               3:
                   IF (("req23" OR "reqdown3") AND "proximity23") THEN
                       #elevator2next := 3;
                   ELSIF ("req22" OR "reqdown2") THEN
                       #elevator2next := 2;
                       #elevator2heading := 1;
                   ELSIF ("req21" OR "reqdown1") THEN
                       #elevator2next := 1;
                       #elevator2heading := 1;
                   ELSIF ("req20") THEN
                       #elevator2next := 0;
                       #elevator2heading := 1;
                   ELSIF ("requpgnd") THEN
                       "requpgnd" := FALSE;
                       "req20" := TRUE;
                       #elevator2next := 0;
                       #elevator2heading := 1;
                   ELSIF ("requp1") THEN
                       "requp1" := FALSE;
                       "req21" := TRUE;
                       #elevator2next := 1;
                       #elevator2heading := 1;
                   ELSIF ("requp2") THEN
                       "requp2" := FALSE;
                       "req22" := TRUE;
                       #elevator2next := 2;
                       #elevator2heading := 1;
                   ELSE
                       #elevator2heading := 0;
                   END_IF;
               4:
                   IF (("req24" OR "reqdown4") AND "proximity24") THEN
                       #elevator2next := 4;
                   ELSIF ("req23" OR "reqdown3") THEN
                       #elevator2next := 3;
                       #elevator2heading := 1;
                   ELSIF ("req22" OR "reqdown2") THEN
                       #elevator2next := 2;
                       #elevator2heading := 1;
                   ELSIF ("req21" OR "reqdown1") THEN
                       #elevator2next := 1;
                       #elevator2heading := 1;
                   ELSIF ("req20") THEN
                       #elevator2next := 0;
                       #elevator2heading := 1;
                   ELSIF ("requpgnd") THEN
                       "requpgnd" := FALSE;
                       "req20" := TRUE;
                       #elevator2next := 0;
                       #elevator2heading := 1;
                   ELSIF ("requp1") THEN
                       "requp1" := FALSE;
                       "req21" := TRUE;
                       #elevator2next := 1;
                       #elevator2heading := 1;
                   ELSIF ("requp2") THEN
                       "requp2" := FALSE;
                       "req22" := TRUE;
                       #elevator2next := 2;
                       #elevator2heading := 1;
                   ELSIF ("requp3") THEN
                       "requp3" := FALSE;
                       "req23" := TRUE;
                       #elevator2next := 3;
                       #elevator2heading := 1;
                   ELSE
                       #elevator2heading := 0;
                   END_IF;

               5:
                   IF (("req25" OR "reqdown5") AND "proximity25") THEN
                       #elevator2next := 5;
                   ELSIF ("req24" OR "reqdown4") THEN
                       #elevator2next := 4;
                       #elevator2heading := 1;
                   ELSIF ("req23" OR "reqdown3") THEN
                       #elevator2next := 3;
                       #elevator2heading := 1;
                   ELSIF ("req22" OR "reqdown2") THEN
                       #elevator2next := 2;
                       #elevator2heading := 1;
                   ELSIF ("req21" OR "reqdown1") THEN
                       #elevator2next := 1;
                       #elevator2heading := 1;
                   ELSIF ("req20") THEN
                       #elevator2next := 0;
                       #elevator2heading := 1;
                   ELSIF ("requpgnd") THEN
                       "requpgnd" := FALSE;
                       "req20" := TRUE;
                       #elevator2next := 0;
                       #elevator2heading := 1;
                   ELSIF ("requp1") THEN
                       "requp1" := FALSE;
                       "req21" := TRUE;
                       #elevator2next := 1;
                       #elevator2heading := 1;
                   ELSIF ("requp2") THEN
                       "requp2" := FALSE;
                       "req22" := TRUE;
                       #elevator2next := 2;
                       #elevator2heading := 1;
                   ELSIF ("requp3") THEN
                       "requp3" := FALSE;
                       "req23" := TRUE;
                       #elevator2next := 3;
                       #elevator2heading := 1;
                   ELSIF ("requp4") THEN
                       "requp4" := FALSE;
                       "req24" := TRUE;
                       #elevator2next := 4;
                       #elevator2heading := 1;

                   ELSE
                       #elevator2heading := 0;
                   END_IF;
           END_CASE;

           ;
       END_IF;

   END_IF;






       IF #elevator1.idling THEN
           CASE "elevator1position" OF
               0:
                   IF ("requpgnd" OR "req10") THEN
                       #elevator1stopidling := TRUE;
                   ELSE
                       #elevator1stopidling := FALSE;
                   END_IF;
                   ;
               1:
                   IF ("requp1" OR "reqdown1" OR "req11") THEN
                       #elevator1stopidling := TRUE;
                   ELSE
                       #elevator1stopidling := FALSE;
                   END_IF;
                   ;
               2:
                   IF ("requp2" OR "reqdown2" OR "req12") THEN
                       #elevator1stopidling := TRUE;
                   ELSE
                       #elevator1stopidling := FALSE;
                   END_IF;
                   ;
               3:
                   IF ("requp3" OR "reqdown3" OR "req13") THEN
                       #elevator1stopidling := TRUE;
                   ELSE
                       #elevator1stopidling := FALSE;
                   END_IF;
                   ;
               4:
                   IF ("requp4" OR "reqdown4" OR "req14") THEN
                       #elevator1stopidling := TRUE;
                   ELSE
                       #elevator1stopidling := FALSE;
                   END_IF;
                   ;
               5:
                   IF ("reqdown5" OR "req15") THEN
                       #elevator1stopidling := TRUE;
                   ELSE
                       #elevator1stopidling := FALSE;
                   END_IF;
                   ;
           END_CASE;

       END_IF;

       IF #elevator2.idling THEN
           CASE "elevator2position" OF
               0:
                   IF ("requpgnd" OR "req20") THEN
                       #elevator2stopidling := TRUE;
                   ELSE
                       #elevator2stopidling := FALSE;
                   END_IF;
                   ;
               1:
                   IF ("requp1" OR "reqdown1" OR "req21") THEN
                       #elevator2stopidling := TRUE;
                   ELSE
                       #elevator2stopidling := FALSE;
                   END_IF;
                   ;
               2:
                   IF ("requp2" OR "reqdown2" OR "req22") THEN
                       #elevator2stopidling := TRUE;
                   ELSE
                       #elevator2stopidling := FALSE;
                   END_IF;
                   ;
               3:
                   IF ("requp3" OR "reqdown3" OR "req23") THEN
                       #elevator2stopidling := TRUE;
                   ELSE
                       #elevator2stopidling := FALSE;
                   END_IF;
                   ;
               4:
                   IF ("requp4" OR "reqdown4" OR "req24") THEN
                       #elevator2stopidling := TRUE;
                   ELSE
                       #elevator2stopidling := FALSE;
                   END_IF;
                   ;
               5:
                   IF ("reqdown5" OR "req25") THEN
                       #elevator2stopidling := TRUE;
                   ELSE
                       #elevator2stopidling := FALSE;
                   END_IF;
                   ;
           END_CASE;

       END_IF;

   #elevator1(currentlevel:="elevator1position",
              doorclosedsens:="door1closedsens",
              dooropensens:="door1opensens",
              nextlevel:=#elevator1next,
              las:=true,
              stopidling:=#elevator1stopidling,
              closethedoorbutton:="doorclosebutton1",
              openthedoorbutton:="dooropenbutton1",
              ack:=#elevator1ack,
              opendoor=>"door1openmotor",
              closedoor=>"door1closemotor",
              headingup=>"elevator1upmotor",
              headingdown=>"elevator1downmotor");
   #elevator2(currentlevel:="elevator2position",
              doorclosedsens:="door2closedsens",
              dooropensens:="door2opensens",
              nextlevel:=#elevator2next,
              las:=TRUE,
              stopidling:=#elevator2stopidling,
              closethedoorbutton:="doorclosebutton2",
              openthedoorbutton:="dooropenbutton2",
              ack:=#elevator2ack,
              opendoor=>"door2openmotor",
              closedoor=>"door2closemotor",
              headingup=>"elevator2upmotor",
              headingdown=>"elevator2downmotor");
END_FUNCTION_BLOCK

FUNCTION "sensors_to_int_position" : Void   // FC1, SCL
{ S7_Optimized_Access := 'TRUE' }
VERSION : 0.1
   VAR_INPUT
      in1g : Bool;
      in11 : Bool;
      in12 : Bool;
      in13 : Bool;
      in14 : Bool;
      in15 : Bool;
      in2g : Bool;
      in21 : Bool;
      in22 : Bool;
      in23 : Bool;
      in24 : Bool;
      in25 : Bool;
   END_VAR
   VAR_OUTPUT
      out1 : Int;
      out2 : Int;
   END_VAR
BEGIN
   IF #in1g THEN
       #out1 := 0;
   END_IF;
   IF #in11 THEN
       #out1 := 1;
   END_IF;
   IF #in12 THEN
       #out1 := 2;
   END_IF;
   IF #in13 THEN
       #out1 := 3;
   END_IF;
   IF #in14 THEN
       #out1 := 4;
   END_IF;
   IF #in15 THEN
       #out1 := 5;
   END_IF;

   IF #in2g THEN
       #out2 := 0;
   END_IF;
   IF #in21 THEN
       #out2 := 1;
   END_IF;
   IF #in22 THEN
       #out2 := 2;
   END_IF;
   IF #in23 THEN
       #out2 := 3;
   END_IF;
   IF #in24 THEN
       #out2 := 4;
   END_IF;
   IF #in25 THEN
       #out2 := 5;
   END_IF;
END_FUNCTION

FUNCTION "input_timers" : Void   // FC2, SCL
{ S7_Optimized_Access := 'TRUE' }
VERSION : 0.1
BEGIN
   "door1closing".TON(IN:="door1closemotor",
                      PT:=T#1s,
                      Q=>"door1closedsens");
   "door1opening".TON(IN:="door1openmotor",
                      PT:=T#1s,
                      Q=>"door1opensens");
   "door2closing".TON(IN:="door2closemotor",
                      PT:=T#1s,
                      Q=>"door2closedsens");
   "door2opening".TON(IN:="door2openmotor",
                      PT:=T#1s,
                      Q=>"door2opensens");


   "starting_up1".TON(IN := (("state1" = 2) AND ("elevator1upmotor")),
                      PT := T#500ms);
   "starting_down1".TON(IN:=(("state1"=3) AND ("elevator1downmotor")),
                        PT:=T#500ms);
   "goingup1".TON(IN:=(("state1"=4) AND ("elevator1upmotor")),
                  PT:=T#5s);
   "goingdown1".TON(IN:=(("state1"=5) AND ("elevator1downmotor")),
                    PT:=T#5s);
   "starting_up2".TON(IN := (("state2" = 2) AND ("elevator2upmotor")),
                      PT := T#500ms);
   "starting_down2".TON(IN:=(("state2"=3) AND ("elevator2downmotor")),
                        PT:=T#500ms);
   "goingup2".TON(IN := (("state2" = 4) AND ("elevator2upmotor")),
                  PT := T#5s);
   "goingdown2".TON(IN:=(("state2"=5) AND ("elevator2downmotor")),
                    PT:=T#5s);


   //states:
   //1:stopped
   //2:start going up
   //3: start going down
   //4: going up
   //5: going down
   //6:arrived up
   //7: arrived down
   //
   CASE "state1" OF
       0:
           "lastfloor1" := 1;
           "state1" := 1;

       1:
           IF "elevator1upmotor" AND (NOT ("proximity15")) THEN
               "state1" := 2;
           ELSIF "elevator1downmotor" AND (NOT ("proximity1ground")) THEN
               "state1" := 3;
           END_IF;

       2:
           IF "starting_up1".Q THEN
               "state1" := 4;
           ELSIF NOT("elevator1upmotor") THEN
               "state1" := 1;
           END_IF;
       3:
           IF "starting_down1".Q THEN
               "state1" := 5;
           ELSIF NOT ("elevator1downmotor") THEN
               "state1" := 1;
           END_IF;
       4:
           IF "goingup1".Q THEN
               "state1" := 6;
           END_IF;
       5:
           IF "goingdown1".Q THEN
               "state1" := 7;
           END_IF;
       6,7:
           "state1" := 1;
       ELSE  // Statement section ELSE
           ;
   END_CASE;

   CASE "state1" OF

       1,2,3:

           "int_to_bools"(in1 := "lastfloor1",
                          out1 => "proximity1ground",
                          out2 => "proximity11",
                          out3 => "proximity12",
                          out4 => "proximity13",
                          out5 => "proximity14",
                          out6 => "proximity15");


       4,5:
           "int_to_bools"(in1 := 0,
                          out1 => "proximity1ground",
                          out2 => "proximity11",
                          out3 => "proximity12",
                          out4 => "proximity13",
                          out5 => "proximity14",
                          out6 => "proximity15");
           ;
       6:
           IF "lastfloor1" < 7 THEN
               "lastfloor1" := "lastfloor1" + 1;
           END_IF;
           "int_to_bools"(in1 := "lastfloor1",
                          out1 => "proximity1ground",
                          out2 => "proximity11",
                          out3 => "proximity12",
                          out4 => "proximity13",
                          out5 => "proximity14",
                          out6 => "proximity15");
       7:
           IF "lastfloor1" > 1 THEN
               "lastfloor1" := "lastfloor1" - 1;
           END_IF;
           "int_to_bools"(in1 := "lastfloor1",
                          out1 => "proximity1ground",
                          out2 => "proximity11",
                          out3 => "proximity12",
                          out4 => "proximity13",
                          out5 => "proximity14",
                          out6 => "proximity15");
       ELSE  // Statement section ELSE
           ;
   END_CASE;

   // second elevator:
   // 
   CASE "state2" OF
       0:
           "lastfloor2" := 1;
           "state2" := 1;

       1:
           IF "elevator2upmotor" AND (NOT ("proximity25")) THEN
               "state2" := 2;
           ELSIF "elevator2downmotor" AND (NOT ("proximity2ground")) THEN
               "state2" := 3;
           END_IF;

       2:
           IF "starting_up2".Q THEN
               "state2" := 4;
           ELSIF NOT("elevator2upmotor") THEN
               "state2" := 1;
           END_IF;
       3:
           IF "starting_down2".Q THEN
               "state2" := 5;
           ELSIF NOT("elevator2downmotor") THEN
               "state2" := 1;
           END_IF;
       4:
           IF "goingup2".Q THEN
               "state2" := 6;
           END_IF;
       5:
           IF "goingdown2".Q THEN
               "state2" := 7;
           END_IF;
       6, 7:
           "state2" := 1;
       ELSE  // Statement section ELSE
           ;
   END_CASE;

   CASE "state2" OF

       1, 2, 3:

           "int_to_bools"(in1 := "lastfloor2",
                          out1 => "proximity2ground",
                          out2 => "proximity21",
                          out3 => "proximity22",
                          out4 => "proximity23",
                          out5 => "proximity24",
                          out6 => "proximity25");


       4, 5:
           "int_to_bools"(in1 := 0,
                          out1 => "proximity2ground",
                          out2 => "proximity21",
                          out3 => "proximity22",
                          out4 => "proximity23",
                          out5 => "proximity24",
                          out6 => "proximity25");
           ;
       6:
           IF "lastfloor2" < 7 THEN
               "lastfloor2" := "lastfloor2" + 1;
           END_IF;
           "int_to_bools"(in1 := "lastfloor2",
                          out1 => "proximity2ground",
                          out2 => "proximity21",
                          out3 => "proximity22",
                          out4 => "proximity23",
                          out5 => "proximity24",
                          out6 => "proximity25");
       7:
           IF "lastfloor2" > 1 THEN
               "lastfloor2" := "lastfloor2" - 1;
           END_IF;
           "int_to_bools"(in1 := "lastfloor2",
                          out1 => "proximity2ground",
                          out2 => "proximity21",
                          out3 => "proximity22",
                          out4 => "proximity23",
                          out5 => "proximity24",
                          out6 => "proximity25");
       ELSE  // Statement section ELSE
           ;
   END_CASE;
END_FUNCTION

FUNCTION "int_to_bools" : Void   // FC3, SCL
{ S7_Optimized_Access := 'TRUE' }
VERSION : 0.1
   VAR_INPUT
      in1 : Int;
   END_VAR
   VAR_OUTPUT
      out1 : Bool;
      out2 : Bool;
      out3 : Bool;
      out4 : Bool;
      out5 : Bool;
      out6 : Bool;
   END_VAR
BEGIN
   CASE #in1 OF
       0:
           #out1 := FALSE;
           #out2 := FALSE;
           #out3 := FALSE;
           #out4 := FALSE;
           #out5 := FALSE;
           #out6 := FALSE;
       1:
           #out1 := TRUE;
           #out2 := FALSE;
           #out3 := FALSE;
           #out4 := FALSE;
           #out5 := FALSE;
           #out6 := FALSE;
       2:
           #out1 := FALSE;
           #out2 := TRUE;
           #out3 := FALSE;
           #out4 := FALSE;
           #out5 := FALSE;
           #out6 := FALSE;
       3:
           #out1 := FALSE;
           #out2 := FALSE;
           #out3 := TRUE;
           #out4 := FALSE;
           #out5 := FALSE;
           #out6 := FALSE;
       4:
           #out1 := FALSE;
           #out2 := FALSE;
           #out3 := FALSE;
           #out4 := TRUE;
           #out5 := FALSE;
           #out6 := FALSE;
       5:
           #out1 := FALSE;
           #out2 := FALSE;
           #out3 := FALSE;
           #out4 := FALSE;
           #out5 := TRUE;
           #out6 := FALSE;
       6:
           #out1 := FALSE;
           #out2 := FALSE;
           #out3 := FALSE;
           #out4 := FALSE;
           #out5 := FALSE;
           #out6 := TRUE;

   END_CASE;
END_FUNCTION

FUNCTION "HMI_doors" : Void   // FC6, SCL
{ S7_Optimized_Access := 'TRUE' }
VERSION : 0.1
BEGIN
   CASE "activefloor" OF
       0:
           IF ("door1opensens" AND "proximity1ground") THEN
               "door1open" := TRUE;
           ELSE
               "door1open" := FALSE;
           END_IF;
           IF ("door2opensens" AND "proximity2ground") THEN
               "door2open" := TRUE;
           ELSE
               "door2open" := FALSE;
           END_IF;
       1:
           IF ("door1opensens" AND "proximity11") THEN
               "door1open" := TRUE;
           ELSE
               "door1open" := FALSE;
           END_IF;
           IF ("door2opensens" AND "proximity21") THEN
               "door2open" := TRUE;
           ELSE
               "door2open" := FALSE;
           END_IF;
       2:
           IF ("door1opensens" AND "proximity12") THEN
               "door1open" := TRUE;
           ELSE
               "door1open" := FALSE;
           END_IF;
           IF ("door2opensens" AND "proximity22") THEN
               "door2open" := TRUE;
           ELSE
               "door2open" := FALSE;
           END_IF;
       3:
           IF ("door1opensens" AND "proximity13") THEN
               "door1open" := TRUE;
           ELSE
               "door1open" := FALSE;
           END_IF;
           IF ("door2opensens" AND "proximity23") THEN
               "door2open" := TRUE;
           ELSE
               "door2open" := FALSE;
           END_IF;
       4:
           IF ("door1opensens" AND "proximity14") THEN
               "door1open" := TRUE;
           ELSE
               "door1open" := FALSE;
           END_IF;
           IF ("door2opensens" AND "proximity24") THEN
               "door2open" := TRUE;
           ELSE
               "door2open" := FALSE;
           END_IF;
       5:
           IF ("door1opensens" AND "proximity15") THEN
               "door1open" := TRUE;
           ELSE
               "door1open" := FALSE;
           END_IF;
           IF ("door2opensens" AND "proximity25") THEN
               "door2open" := TRUE;
           ELSE
               "door2open" := FALSE;
           END_IF;
   END_CASE;
END_FUNCTION

ORGANIZATION_BLOCK "Main"   // OB1, LAD, ProgramCycle
TITLE = "Main Program Sweep (Cycle)"
{ S7_Optimized_Access := 'TRUE' }
VERSION : 0.1
BEGIN
END_ORGANIZATION_BLOCK

ORGANIZATION_BLOCK "Simulation"   // OB123, LAD, ProgramCycle
TITLE = "Main Program Sweep (Cycle)"
{ S7_Optimized_Access := 'TRUE' }
VERSION : 0.1
BEGIN
END_ORGANIZATION_BLOCK

(* ===== HMI "HMI_RT_1" =====
system functions are stored by id; their names below are inferred from use
connection "HMI_Connection_1": ETHERNET, SMART_S7_1200_OMS

HMI tags "Default tag table"
   "Tag_ScreenNumber" : UInt, internal
   "elevator1location" : Int = PLC elevator1position AT %MW28, 1 s
   "elevator2location" : Int = PLC elevator2position AT %MW26, 1 s
   "elevator1heading" : Int = PLC ControlBlock_DB.elevator1heading AT %DB1.DBW0, 1 s
   "elevator2heading" : Int = PLC ControlBlock_DB.elevator2heading AT %DB1.DBW0, 1 s
   "activefloor" : Int = PLC activefloor AT %MW40, 1 s
   "door1open" : Bool = PLC door1open AT %M42.0, 1 s
   "door2open" : Bool = PLC door2open AT %M42.1, 1 s
   "elevator1downmotor" : Bool = PLC elevator1downmotor AT %M9.1, 1 s
   "elevator2upmotor" : Bool = PLC elevator2upmotor AT %M9.2, 1 s
   "elevator2downmotor" : Bool = PLC elevator2downmotor AT %M9.3, 1 s
   "elevator1upmotor" : Bool = PLC elevator1upmotor AT %M9.0, 1 s
   "door1opensens" : Bool = PLC door1opensens AT %M8.2, 1 s
   "door1closedsens" : Bool = PLC door1closedsens AT %M8.3, 1 s
   "door2opensens" : Bool = PLC door2opensens AT %M8.4, 1 s

HMI tags "Liftinside"
   "req10" : Bool = PLC req10 AT %M4.2, 1 s
   "req11" : Bool = PLC req11 AT %M4.3, 1 s
   "req12" : Bool = PLC req12 AT %M4.4, 1 s
   "req13" : Bool = PLC req13 AT %M4.5, 1 s
   "req14" : Bool = PLC req14 AT %M4.6, 1 s
   "req15" : Bool = PLC req15 AT %M4.7, 1 s
   "req20" : Bool = PLC req20 AT %M5.0, 1 s
   "req21" : Bool = PLC req21 AT %M5.1, 1 s
   "req22" : Bool = PLC req22 AT %M5.2, 1 s
   "req23" : Bool = PLC req23 AT %M5.3, 1 s
   "req24" : Bool = PLC req24 AT %M5.4, 1 s
   "req25" : Bool = PLC req25 AT %M5.5, 1 s
   "requpgnd" : Bool = PLC requpgnd AT %M7.0, 1 s
   "requp1" : Bool = PLC requp1 AT %M7.1, 1 s
   "requp2" : Bool = PLC requp2 AT %M7.2, 1 s
   "requp3" : Bool = PLC requp3 AT %M7.3, 1 s
   "requp4" : Bool = PLC requp4 AT %M7.4, 1 s
   "reqdown5" : Bool = PLC reqdown5 AT %M7.5, 1 s
   "reqdown4" : Bool = PLC reqdown4 AT %M7.6, 1 s
   "reqdown3" : Bool = PLC reqdown3 AT %M7.7, 1 s
   "reqdown2" : Bool = PLC reqdown2 AT %M5.6, 1 s
   "reqdown1" : Bool = PLC reqdown1 AT %M5.7, 1 s
   "las2" : Bool = PLC las2 AT %M6.1, 1 s
   "las1" : Bool = PLC las1 AT %M6.0, 1 s
   "doorclosebutton1" : Bool = PLC doorclosebutton1 AT %M6.2, 1 s
   "doorclosebutton2" : Bool = PLC doorclosebutton2 AT %M6.3, 1 s
   "dooropenbutton1" : Bool = PLC dooropenbutton1 AT %M6.4, 1 s
   "dooropenbutton2" : Bool = PLC dooropenbutton2 AT %M6.5, 1 s

text list "floors": 0 'Ground Floor'; 1 '1st Floor'; 2 '2nd Floor'; 3 '3rd Floor'; 4 '4th Floor'; 5 '5th Floor'

Template "elevatortemplate" 800x480
   Button "Template_Button" at 614,429 size 71x50; TextOff 'Text'
   Button "Template_Button_1" at 514,429 size 71x50; TextOff 'Text'
   Button "Template_Button_2" at 414,429 size 71x50; TextOff 'Text'
   Button "Template_Button_3" at 314,429 size 71x50; TextOff 'Text'
   Button "Template_Button_4" at 214,429 size 71x50; TextOff 'KÜLSŐ'
      on Release: ActivateScreen("floor1", 0)
   DateTimeField "HmiScreenItemData" at 695,25 size 105x25
   DateTimeField "HmiScreenItemData_1" at 695,0 size 105x25
   Button "Template_Button_6" at 114,429 size 71x50; TextOff 'LIFT2'
      on Release: ActivateScreen("Elevator2 Inside Panel", 0)
   Button "Template_Button_7" at 14,429 size 71x50; TextOff 'LIFT1'
      on Release: ActivateScreen("Elevator1 Inside Panel", 0)
   Button "Template_Button_8" at 714,429 size 71x50; TextOff 'Text'

screen "Root screen" 800x480, template "elevatortemplate"
   on GenerateScreen: SetTag("Tag_ScreenNumber", 1)
   TextField "HmiScreenItemData" at 80,225 size 640x25; Text 'Welcome to KTP700.Basic (KTP700 Basic+ PN)!'
   Button "HmiScreenItemData_1" at 36,87 size 159x47; TextOff 'SIMATIC PLC system diagnos...'; PictureOff "Navigates to SIMATIC PLC system diagnostics for KTP700 Basic+ PN 17.0.0.0"; PictureOn "Navigates to SIMATIC PLC system diagnostics for KTP700 Basic+ PN 17.0.0.0"
      on Release: ActivateScreen("SIMATIC PLC system diagnostics", 0)
   Button "HmiScreenItemData_2" at 36,146 size 159x47; TextOff 'Project information'; PictureOff "Navigates to Project information for KTP700 Basic+ PN 17.0.0.0"; PictureOn "Navigates to Project information for KTP700 Basic+ PN 17.0.0.0"
      on Release: ActivateScreen("Project information", 0)
   Button "HmiScreenItemData_3" at 36,205 size 159x47; TextOff 'User administration'; PictureOff "Navigates to User administration for KTP700 Basic+ PN 17.0.0.0"; PictureOn "Navigates to User administration for KTP700 Basic+ PN 17.0.0.0"
      on Release: ActivateScreen("User administration", 0)
   Button "HmiScreenItemData_4" at 36,264 size 159x47; TextOff 'System information'; PictureOff "Navigates to System information for KTP700 Basic+ PN 17.0.0.0"; PictureOn "Navigates to System information for KTP700 Basic+ PN 17.0.0.0"
      on Release: ActivateScreen("System information", 0)
   Button "HmiScreenItemData_5" at 36,323 size 159x47; TextOff 'Different jobs'; PictureOff "Navigates to Different jobs for KTP700 Basic+ PN 17.0.0.0"; PictureOn "Navigates to Different jobs for KTP700 Basic+ PN 17.0.0.0"
      on Release: ActivateScreen("Different jobs", 0)

screen "SIMATIC PLC system diagnostics" 800x480, template "elevatortemplate"
   on GenerateScreen: SetTag("Tag_ScreenNumber", 2)
   SysDiagControl "HmiScreenItemData" at 1,100 size 796x321
   Button "Back" at 1,52 size 159x47; TextOff 'Back'
      on Release: ActivateScreen("Root screen", 0)

screen "Project information" 800x480, template "elevatortemplate"
   on GenerateScreen: SetTag("Tag_ScreenNumber", 3)
   TextField "HmiScreenItemData" at 35,102 size 171x28; Text 'Project name:'
   TextField "HmiScreenItemData_1" at 241,102 size 524x28; Text 'AUTdevices'
   TextField "HmiScreenItemData_2" at 35,132 size 171x28; Text 'Created on:'
   TextField "HmiScreenItemData_3" at 241,132 size 524x28; Text '3/11/2024 9:57:34 AM'
   TextField "HmiScreenItemData_4" at 35,162 size 171x28; Text 'Author:'
   TextField "HmiScreenItemData_5" at 241,162 size 524x28; Text 'PLCDev'
   TextField "HmiScreenItemData_6" at 35,192 size 171x28; Text 'Description:'
   TextField "HmiScreenItemData_7" at 241,192 size 524x28; Text 'Az Automatizálási Tanszék SIMATIC eszközei'
   Button "Back" at 1,52 size 159x47; TextOff 'Back'
      on Release: ActivateScreen("Root screen", 0)

screen "User administration" 800x480, template "elevatortemplate"
   on GenerateScreen: SetTag("Tag_ScreenNumber", 4)
   UserView "HmiScreenItemData" at 1,100 size 796x321
   Button "Back" at 1,52 size 159x47; TextOff 'Back'
      on Release: ActivateScreen("Root screen", 0)

screen "System information" 800x480, template "elevatortemplate"
   on GenerateScreen: SetTag("Tag_ScreenNumber", 5)
   TextField "HmiScreenItemData" at 35,102 size 171x28; Text 'HMI device type:'
   TextField "HmiScreenItemData_1" at 241,102 size 524x28; Text 'KTP700 Basic+ PN 17.0.0.0'
   TextField "HmiScreenItemData_2" at 35,132 size 171x28; Text 'Connection:'
   TextField "HmiScreenItemData_3" at 241,132 size 524x28; Text 'PROFINET (X1)'
   TextField "HmiScreenItemData_4" at 35,162 size 171x28; Text 'PLC:'
   TextField "HmiScreenItemData_5" at 241,162 size 524x28; Text 'SIMATIC S7 1200'
   Button "Back" at 1,52 size 159x47; TextOff 'Back'
      on Release: ActivateScreen("Root screen", 0)

screen "Different jobs" 800x480, template "elevatortemplate"
   on GenerateScreen: SetTag("Tag_ScreenNumber", 6)
   Button "Online" at 36,146 size 159x47; TextOff 'Online'
      on Release: function_bb44b551(0)
   Button "Offline" at 36,205 size 159x47; TextOff 'Offline'
      on Release: function_bb44b551(1)
   Button "Transfer" at 36,264 size 159x47; TextOff 'Transfer'
      on Release: function_bb44b551(2)
   Button "Toggle language" at 36,323 size 159x47; TextOff 'Toggle language'
      on Release: function_fb9197e8(-1)
   Button "Stop Runtime" at 207,146 size 159x47; TextOff 'Stop Runtime'
      on Release: StopRuntime(0)
   Button "Back" at 1,52 size 159x47; TextOff 'Back'
      on Release: ActivateScreen("Root screen", 0)

screen "Elevator1 Inside Panel" 800x480, template "elevatortemplate"
   on GenerateScreen: SetTag("Tag_ScreenNumber", 4)
   Button "Button_1" at 470,62 size 58x59; TextOff '4'
      on Click: SetBit("req14")
   Button "Button_2" at 577,62 size 58x59; TextOff '5'
      on Click: SetBit("req15")
   Button "Button_3" at 470,149 size 58x59; TextOff '2'
      on Click: SetBit("req12")
   Button "Button_4" at 577,149 size 58x59; TextOff '3'
      on Click: SetBit("req13")
   Button "Button_5" at 577,235 size 58x59; TextOff '1'
      on Click: SetBit("req11")
   Button "Button_6" at 470,235 size 58x59; TextOff '0'
      on Click: SetBit("req10")
   Button "Button_7" at 472,320 size 58x59; TextOff 'Text'
      on Press: SetBit("dooropenbutton1")
      on Release: ResetBit("dooropenbutton1")
   Button "Button_8" at 577,320 size 58x59; TextOff 'Text'
      on Press: SetBit("doorclosebutton1")
      on Release: ResetBit("doorclosebutton1")
   GraphicView "elevator1closed" at 70,59 size 273x349; Picture "doorclosed1"
      Visibility <- "door1opensens"
   GraphicView "elevator1open" at 70,58 size 273x350; Picture "dooropened1"
      Visibility <- "door1opensens"
   GraphicView "elevator1idleindicator" at 167,15 size 76x33; Picture "idle"
   GraphicView "Graphic view_1" at 417,25 size 274x394; Picture "elevatorpanel"
   TextField "Text field_1" at 517,28 size 75x33; Text 'LIFT1'
   GraphicView "elevator1upindicator" at 167,15 size 76x33; Picture "headingup"
      Visibility <- "elevator1upmotor"
   GraphicView "elevator1downindicator" at 168,15 size 77x33; Picture "headingdown"
      Visibility <- "elevator1downmotor"
   IOField "I/O field_1" at 200,14 size 38x32; FormatPattern 9
      ProcessValue <- "elevator1location"

Template "defaulttemplate" 800x480
   Button "Exit" at 714,429 size 71x50; TextOn 'Exit'; TextOff 'Exit'; PictureOn "ExitRuntime_KTP700_Basic_PN_TR"; PictureOff "ExitRuntime_KTP700_Basic_PN_TR"
      on Release: StopRuntime(0)
   Button "Template_Button" at 614,429 size 71x50; TextOff 'Text'
   Button "Template_Button_1" at 514,429 size 71x50; TextOff 'Text'
   Button "Template_Button_2" at 414,429 size 71x50; TextOff 'Text'
   Button "Template_Button_3" at 314,429 size 71x50; TextOff 'Text'
   Button "Template_Button_4" at 214,429 size 71x50; TextOff 'Text'
   Button "Alarms" at 114,429 size 71x50; TextOn 'Alarms'; TextOff 'Alarms'; PictureOn "AlarmDisplay_KTP700_Basic_PN_TR"; PictureOff "AlarmDisplay_KTP700_Basic_PN_TR"
      on Release: function_ef3f5d25("Alarm window_Unacknowledged", -1)
   Button "Start screen" at 14,429 size 71x50; TextOn 'Start screen'; TextOff 'Start screen'; PictureOn "NavigateHome_KTP700_Basic_PN_TR"; PictureOff "NavigateHome_KTP700_Basic_PN_TR"
      on Release: ActivateScreen("Elevator1 Inside Panel", 7)
   SymbolicIOField "Symbolic_IO_Field_Screen" at 93,9 size 600x33; TextOn '1'; TextOff '0'; TextList "TextList_ScreenNames"
      on Change: ActivateScreenByNumber("Tag_ScreenNumber", 0)
      ProcessValue <- "Tag_ScreenNumber"
   DateTimeField "HmiScreenItemData" at 695,25 size 105x25
   DateTimeField "HmiScreenItemData_1" at 695,0 size 105x25
   GraphicView "Logo" at 0,0 size 91x51; Picture "Logo of KTP700.Basic"

screen "Elevator2 Inside Panel" 800x480, template "elevatortemplate"
   GraphicView "Graphic view_1" at 417,25 size 274x394; Picture "elevatorpanel"
   TextField "Text field_1" at 517,28 size 75x33; Text 'LIFT2'
   Button "Button_1" at 470,62 size 58x59; TextOff '4'
      on Click: SetBit("req24")
   Button "Button_2" at 577,62 size 58x59; TextOff '5'
      on Click: SetBit("req25")
   Button "Button_3" at 470,149 size 58x59; TextOff '2'
      on Click: SetBit("req22")
   Button "Button_4" at 577,149 size 58x59; TextOff '3'
      on Click: SetBit("req23")
   Button "Button_5" at 577,235 size 58x59; TextOff '1'
      on Click: SetBit("req21")
   Button "Button_6" at 470,235 size 58x59; TextOff '0'
      on Click: SetBit("req20")
   Button "Button_7" at 472,320 size 58x59; TextOff 'Text'
      on Release: ResetBit("dooropenbutton2")
      on Press: SetBit("dooropenbutton2")
   Button "Button_8" at 577,320 size 58x59; TextOff 'Text'
      on Release: ResetBit("doorclosebutton2")
      on Press: SetBit("doorclosebutton2")
   GraphicView "elevator2open" at 70,55 size 273x350; Picture "dooropened1"
      Visibility <- "door2opensens"
   GraphicView "elevator2closed" at 70,56 size 273x358; Picture "doorclosed1"
      Visibility <- "door2opensens"
   GraphicView "elevator2idleindicator" at 168,16 size 76x33; Picture "idle"
   GraphicView "elevator2upindicator" at 169,15 size 76x33; Picture "headingup"
      Visibility <- "elevator2upmotor"
   GraphicView "elevator2downindicator" at 168,15 size 77x33; Picture "headingdown"
      Visibility <- "elevator2downmotor"
   IOField "I/O field_3" at 197,15 size 38x32; FormatPattern 9
      ProcessValue <- "elevator2location"

screen "floor1" 800x480, template "elevatortemplate"
   GraphicView "elevator2open" at 501,61 size 273x350; Picture "dooropened1"
      Visibility <- "door2open"
   GraphicView "requestpanel" at 350,136 size 100x200; Picture "istockphoto-1288408696-612x612"
      Visibility <- "activefloor"
   GraphicView "elevator1closed" at 25,62 size 273x349; Picture "doorclosed1"
      Visibility <- "door1open"
   GraphicView "elevator1open" at 25,61 size 273x350; Picture "dooropened1"
      Visibility <- "door1open"
   GraphicView "elevator2closed" at 501,62 size 273x358; Picture "doorclosed1"
      Visibility <- "door2open"
   GraphicView "elevator1idleindicator" at 122,18 size 76x33; Picture "idle"
   GraphicView "elevator2idleindicator" at 599,22 size 76x33; Picture "idle"
   SymbolicIOField "floorselector" at 325,32 size 152x32; TextOff '0'; TextOn '1'; TextList "floors"
      ProcessValue <- "activefloor"
   GraphicView "elevator1upindicator" at 122,18 size 76x33; Picture "headingup"
      Visibility <- "elevator1upmotor"
   GraphicView "elevator1downindicator" at 123,18 size 77x33; Picture "headingdown"
      Visibility <- "elevator1downmotor"
   GraphicView "elevator2upindicator" at 600,21 size 76x33; Picture "headingup"
      Visibility <- "elevator2upmotor"
   GraphicView "elevator2downindicator" at 599,21 size 77x33; Picture "headingdown"
      Visibility <- "elevator2downmotor"
   Button "floor1up" at 368,159 size 65x70; TextOff 'Text'
      on Release: SetTag("requp1", 1)
      Visibility <- "activefloor"
   Button "floor1down" at 370,246 size 65x70; TextOff 'Text'
      on Release: SetTag("reqdown1", 1)
      Visibility <- "activefloor"
   Button "floor2up" at 370,159 size 65x70; TextOff 'Text'
      on Release: SetTag("requp2", 1)
      Visibility <- "activefloor"
   Button "floor2down" at 366,246 size 65x70; TextOff 'Text'
      on Release: SetTag("reqdown2", 1)
      Visibility <- "activefloor"
   Button "floor3down" at 368,246 size 65x70; TextOff 'Text'
      on Release: SetTag("reqdown3", 1)
      Visibility <- "activefloor"
   Button "floor3up" at 370,159 size 65x70; TextOff 'Text'
      on Release: SetTag("requp3", 1)
      Visibility <- "activefloor"
   Button "floor4up" at 366,159 size 65x70; TextOff 'Text'
      on Release: SetTag("requp4", 1)
      Visibility <- "activefloor"
   Button "floor4down" at 370,247 size 65x70; TextOff 'Text'
      on Release: SetTag("reqdown4", 1)
      Visibility <- "activefloor"
   Button "floor5down" at 368,200 size 65x70; TextOff 'Text'
      on Release: SetTag("reqdown5", 1)
      Visibility <- "activefloor"
   Button "floor0up" at 368,200 size 65x70; TextOff 'Text'
      on Release: SetTag("requpgnd", 1)
      Visibility <- "activefloor"
   IOField "I/O field_1" at 155,17 size 38x32; FormatPattern 9
      ProcessValue <- "elevator1location"
   IOField "I/O field_3" at 628,21 size 38x32; FormatPattern 9
      ProcessValue <- "elevator2location"
   GraphicView "groundfloorbutton" at 350,187 size 100x100; Picture "downbutton"
      Visibility <- "activefloor"
   GraphicView "topfloorbutton" at 350,187 size 100x100; Picture "upbutton"
      Visibility <- "activefloor"
*)